(* Logix 5000 project; controller PLC_MCC1300_75F1 vendor 1 type 14 code 166 rev 32.11; software revision 32.04; part 78 of 83 *)
(* tags used below, declared in another part *)
   CM_AreaStackerToLine_JS1_Sync : CM_AreaStackerToLine;
   CM_ConveyorStackerToLine_JS1_Sync : CM_ConveyorStackerToLine;
   M310B : MAC_Conveyor;
   M310B_ALM : MAC_Conveyor_ALM;
   M310B_HMW : MAC_Conveyor_HMW;
   M310Popup : MAC_Popup_ZC[2];
   M311 : MAC_Conveyor;
   M311_ALM : MAC_Conveyor_ALM;
   M311_HMW : MAC_Conveyor_HMW;
   M311A : MAC_Rotator;
   M311A_ALM : MAC_Rotator_ALM;
   M312 : MAC_Conveyor_Single;
   M312_ALM : MAC_Conveyor_ALM;
   M312_HMW : MAC_Conveyor_HMW;
   M350Popup : MAC_Popup_ZC;
   M351 : MAC_Conveyor;
   M351_HMW : MAC_Conveyor_HMW;
   M352 : MAC_Conveyor;
   M352_HMW : MAC_Conveyor_HMW;
   M353 : MAC_Conveyor;
   M353_HMW : MAC_Conveyor_HMW;
   xAlwaysOFF : BOOL;
   xAlwaysON : BOOL;
   Z301 : MAC_Zone_ML;
   Z401 : MAC_Zone;
   Z401_HMR : MAC_Zone_HMR;
   Z401_HMW : MAC_Zone_HMW;
   Z402 : MAC_Zone;
   Z402_ALM : MAC_Zone_ALM;
   Z402_HMR : MAC_Zone_HMR;
   Z402_HMW : MAC_Zone_HMW;
   Z402_INPUT_xMainLineEmergencyON : BOOL;
   Z402_OUTPUT_xMCC_SafetyPanel1 : BOOL;
   Z900 : MAC_Zone;
   Z900_ALM : MAC_Zone_ALM;
   Z900_HMR : MAC_Zone_HMR;
   Z900_HMW : MAC_Zone_HMW;
(* MainProgram, continued *)

   42: [XIC(Z401_HMW.rgxMan.0) OTE(Z401_HMR.rgxMan.0) ,XIC(Z401_HMW.rgxMan.1) OTE(Z401_HMR.rgxMan.1) ];
END_ROUTINE

ROUTINE Z402_Alarm   (* ladder *)
   0: XIC(Z401.tmON_ResetAlarm.DN)FLL(0,Z402_ALM,1);
END_ROUTINE

ROUTINE Z402_Logic   (* ladder *)
   // #####_COSTANTS_#####
   0: NOP();
   // #####_MATCH_#####
   1: NOP();
   // #####_ALARMS_#####
   2: NOP();
   3: XIC(Z402_HMW.xResetErrorRequest)[OTU(Z402_HMW.xResetErrorRequest) ,TOF(Z402.tmON_ResetAlarm,?,?) ];
   4: XIC(Z402.tmON_24Vdc.DN)XIC(Z402.tmON_400Vca.DN)XIC(Z402.tmON_EmergencyOK.DN)OTE(Z402.ST_xEnableControlError);
   5: JSR(Z402_Alarm,0);
   // #####_HMI_LOGICS_#####
   6: NOP();
   // #####_STATUSES_#####
   7: NOP();
   8: [NEQ(Z402_ALM.rgxEmergency[0],0) ,NEQ(Z402_ALM.rgxFault[0],0) ,NEQ(Z402_ALM.rgxWarning[0],0) ,XIC(M310Popup[0].ST_xMachineAlarm) ,XIC(M310Popup[1].ST_xMachineAlarm) ,XIC(M311.ST_xMachineAlarm) ,XIC(M311A.ST_xMachineAlarm) ,XIC(M312.ST_xMachineAlarm) ]OTE(Z402.ST_xZoneError);
   // #####_ZONE MODALITY_#####
   9: NOP();
   // Selector manual mode
   10: XIC(Z402_HMW.xManualModeRequest)OTL(Z402.ST_xSelectionManualMode)OTU(Z402.ST_xSelectionAutomaticMode)OTU(Z402_HMW.xManualModeRequest);
   // Selector automatic mode
   11: XIC(Z402_HMW.xAutomaticModeRequest)OTL(Z402.ST_xSelectionAutomaticMode)OTU(Z402.ST_xSelectionManualMode)OTU(Z402_HMW.xAutomaticModeRequest);
   // Condition Ok for manual mode
   12: [XIC(Z402.ST_xConditionOKStopCycle) ,XIO(Z402.ST_xCycleON) ]OTE(Z402.ST_xConditionOkManualMode);
   // Manual mode accepted
   13: XIC(Z402.ST_xSelectionManualMode)[XIO(Z402.ST_xManualModeAccepted) OTE(Z402.ST_xManualModeRequest) ,[XIC(Z402.ST_xConditionOkManualMode) ,XIC(Z402.ST_xManualModeAccepted) ] OTE(Z402.ST_xManualModeAccepted) ];
   // Auto mode accepted
   14: XIO(Z402.ST_xManualModeAccepted)[XIC(Z402.ST_xSelectionAutomaticMode) ,XIC(Z402.ST_xAutoModeAccepted) ][OTE(Z402.ST_xAutoModeAccepted) ,ONS(Z402.OSR_xAutomaticMode) OTE(Z402.OS_xAutomaticMode) ];
   // Set all manual command for iFix
   15: XIC(Z402.ST_xManualModeAccepted)OTL(M310B_HMW.xEnableDisableManualCommand)OTL(M311_HMW.xEnableDisableManualCommand)OTL(M312_HMW.xEnableDisableManualCommand);
   // Reset all manual command for iFix
   16: XIC(Z402.OS_xAutomaticMode)OTU(M310B_HMW.xEnableDisableManualCommand)OTU(M311_HMW.xEnableDisableManualCommand)OTU(M312_HMW.xEnableDisableManualCommand);
   // #####_LOGICS_#####
   17: NOP();
   18: [XIC(Z402_HMW.xStartCycleRequest) ,XIC(CM_AreaStackerToLine_JS1_Sync.xSB_LineCycle) ]OTE(Z402.OS_xStartCycle);
   19: [XIC(Z402_HMW.xStopCycleRequest) ,XIC(CM_AreaStackerToLine_JS1_Sync.xSB_StopLineCycle) ]OTE(Z402.OS_xStopCycle);
   20: [XIC(Z402.tmON_ForceStop.DN) ONS(Z402.OSR_xForceStopCycle) ,XIC(Z402_HMW.xForceStopCycle) ]OTE(Z402.OS_xForceStopCycle);
   21: XIO(Z402.OS_xForceStopCycle)XIC(Z402.tmON_24Vdc.DN)XIC(Z402.tmON_400Vca.DN)XIC(Z402.tmON_EmergencyOK.DN)OTE(Z402.ST_xConditionOkCycleON);
   22: [XIC(Z402.OS_xStartCycle) ,XIC(Z402.ST_xStartCycleRequest) ]XIC(Z402.ST_xConditionOkCycleON)XIO(Z402.ST_xCycleON)XIO(Z402.OS_xStopCycle)OTE(Z402.ST_xStartCycleRequest);
   23: [XIC(Z402.OS_xStopCycle) ,XIC(Z402.ST_xStopCycleRequest) ]XIC(Z402.ST_xCycleON)XIO(Z402.ST_xStartCycleRequest)OTE(Z402.ST_xStopCycleRequest);
   24: XIC(M310B.ST_xConditionOKStopCycle)XIC(M311.ST_xConditionOKStopCycle)XIC(M311A.ST_xConditionOKStopCycle)XIC(M312.ST_xConditionOKStopCycle)XIC(CM_ConveyorStackerToLine_JS1_Sync.xConditionOkForStopCycle)OTE(Z402.ST_xConditionOKStopCycle);
   25: [XIC(Z402.ST_xStopCycleRequest) XIC(Z402.ST_xConditionOKStopCycle) ,XIC(Z402_HMW.xForceStopCycle) ]OTE(Z402.ST_xStopCycleAccepted);
   // Reimpostare tempo a 15 secondi
   26: [XIC(Z402.ST_xStartCycleRequest) ,XIC(Z402.ST_xCycleON) ]XIC(Z402.ST_xConditionOkCycleON)XIO(Z402.ST_xStopCycleAccepted)XIO(Z402.ST_xManualModeAccepted)[TON(Z402.tmON_Cycle,?,?) ,XIC(Z402.tmON_Cycle.DN) OTE(Z402.ST_xCycleON) ];
   27: XIC(Z402.ST_xCycleON)XIO(Z402.ST_xManualModeRequest)XIO(Z402.ST_xStopCycleRequest)OTE(Z402.ST_xConditionOkPhaseAdvancement);
   28: XIC(Z402.ST_xCycleON)[XIC(M310B.ST_xCleaningAccepted) ,XIO(M310B.ST_xReqCleaning) ][XIC(M311.ST_xCleaningAccepted) ,XIO(M311.ST_xReqCleaning) ][XIC(M312.ST_xCleaningAccepted) ,XIO(M312.ST_xReqCleaning) ]OTE(Z402.ST_xCleaningConditionOK);
   // Speed manager
   29: [MOV(Z402_HMW.dLineSpeed_mm_min,Z402_HMR.dLineSpeed_mm_min) ,LES(Z402_HMR.dLineSpeed_mm_min,35000) MOV(35000,Z402_HMR.dLineSpeed_mm_min) ,GRT(Z402_HMR.dLineSpeed_mm_min,60000) MOV(60000,Z402_HMR.dLineSpeed_mm_min) ];
   // #####_CLEANING_#####
   30: NOP();
   31: XIO(Z402.ST_xCleaningAccepted)XIC(Z402_HMW.xStartCleanZoneRequest)[MOV(Z402_HMW.dCleaningSelection,Z402_HMR.dCleaningSelection) ,OTL(Z402.ST_xReqCleaning) ];
   32: XIC(Z402.ST_xReqCleaning)XIC(Z402.ST_xCleaningConditionOK)[OTL(Z402.ST_xCleaningAccepted) ,OTU(Z402.ST_xReqCleaning) ,OTL(M310B_HMW.xLocalCleaningRequest) ,OTL(M311_HMW.xLocalCleaningRequest) ,OTL(M312_HMW.xLocalCleaningRequest) ];
   33: XIC(Z402_HMW.xStopCleanZoneRequest)[OTU(Z402.ST_xReqCleaning) ,OTU(Z402.ST_xCleaningAccepted) ,MOV(0,Z402_HMW.dCleaningSelection) ,OTU(M310B_HMW.xLocalCleaningRequest) ,OTU(M311_HMW.xLocalCleaningRequest) ,OTU(M311_HMW.xLocalCleaningRequest) ];
   34: XIC(xAlwaysON)[OTU(Z402_HMW.xStartCycleRequest) ,OTU(Z402_HMW.xStopCycleRequest) ,OTU(Z402_HMW.xStartCleanZoneRequest) ,OTU(Z402_HMW.xForceStopCycle) ,OTU(Z402_HMW.xStopCleanZoneRequest) ];
   // #####_HMI_STATUSES_#####
   35: NOP();
   36: XIC(Z402.ST_xZoneError)OTE(Z402_HMR.xZoneAlarm);
   37: [XIC(Z402.ST_xCleaningAccepted) ,XIC(M310B.ST_xCleaningAccepted) XIC(M311.ST_xCleaningAccepted) XIC(M312.ST_xCleaningAccepted) ]OTE(Z402_HMR.xCleaningEnabled);
   38: [MOV(0,Z402_HMR.dCabinetState1) ,[XIC(M310B_ALM.rgxStoppingFault_M[0].1) ,XIC(M311_ALM.rgxStoppingFault_M[0].1) ,XIC(M311A_ALM.rgxStoppingFault_M[0].1) ,XIC(M312_ALM.rgxStoppingFault_M[0].1) ] MOV(2,Z402_HMR.dCabinetState1) ,XIC(Z402_OUTPUT_xMCC_SafetyPanel1) MOV(1,Z402_HMR.dCabinetState1) ];
   39: [XIC(Z402.ST_xManualModeAccepted) MOV(1,Z402_HMR.dZoneMode) ,XIC(Z402.ST_xAutoModeAccepted) MOV(4,Z402_HMR.dZoneMode) ,XIC(Z402.ST_xManualModeRequest) MOV(8,Z402_HMR.dZoneMode) ];
   40: [MOV(2,Z402_HMR.dZoneState) ,XIC(Z402.ST_xStartCycleRequest) XIO(Z402.ST_xCycleON) MOV(4,Z402_HMR.dZoneState) ,XIC(Z402.ST_xCycleON) MOV(1,Z402_HMR.dZoneState) ,XIC(Z402.ST_xStopCycleRequest) MOV(8,Z402_HMR.dZoneState) ,XIO(Z402_INPUT_xMainLineEmergencyON) MOV(1024,Z402_HMR.dZoneState) ];
   41: [[XIC(Z402.ST_xCleaningAccepted) ,XIC(M310B.ST_xCleaningAccepted) XIC(M311.ST_xCleaningAccepted) XIC(M312.ST_xCleaningAccepted) ] MOV(1,Z402_HMR.dCleaningState) ,XIO(Z402.ST_xCleaningAccepted) MOV(2,Z402_HMR.dCleaningState) ,XIC(Z402.ST_xReqCleaning) XIO(Z402.ST_xCleaningAccepted) MOV(4,Z402_HMR.dCleaningState) ];
   42: [XIC(Z402_HMW.rgxMan.0) OTE(Z402_HMR.rgxMan.0) ,XIC(Z402_HMW.rgxMan.1) OTE(Z402_HMR.rgxMan.1) ];
END_ROUTINE

ROUTINE Z900_Alarm   (* ladder *)
   0: XIC(Z900.tmON_ResetAlarm.DN)FLL(0,Z900_ALM,1);
END_ROUTINE

ROUTINE Z900_Logic   (* ladder *)
   // #####_COSTANTS_#####
   0: NOP();
   // #####_MATCH_#####
   1: NOP();
   2: XIC(Z301.INPUT_x24VdcVoltageON)XIC(Z301.INPUT_xPowerSupply24VLogic1)XIC(Z301.INPUT_xPowerSupply24VLogic2)XIC(Z301.INPUT_xPowerSupply24VLogic3)XIC(Z301.INPUT_xEthernetSwitch24VON)XIC(Z301.INPUT_xPowerSupply24VDrive1)XIC(Z301.INPUT_xPowerSupply24VDrive2)TON(Z900.tmON_24Vdc,?,?);
   3: XIC(Z301.INPUT_xPowerSupply400VDrive1)XIC(Z301.INPUT_xPowerSupply400VDrive2)TON(Z900.tmON_400Vca,?,?);
   4: XIC(Z301.INPUT_xMainEmergencyON)TON(Z900.tmON_EmergencyOK,?,?);
   // #####_ALARMS_#####
   5: NOP();
   6: XIC(Z900_HMW.xResetErrorRequest)[OTU(Z900_HMW.xResetErrorRequest) ,TOF(Z900.tmON_ResetAlarm,?,?) ];
   7: XIC(Z900.tmON_24Vdc.DN)XIC(Z900.tmON_400Vca.DN)XIC(Z900.tmON_EmergencyOK.DN)OTE(Z900.ST_xEnableControlError);
   8: JSR(Z900_Alarm,0);
   // #####_HMI_LOGICS_#####
   9: NOP();
   // #####_STATUSES_#####
   10: NOP();
   11: [NEQ(Z900_ALM.rgxEmergency[0],0) ,NEQ(Z900_ALM.rgxFault[0],0) ,NEQ(Z900_ALM.rgxWarning[0],0) ,XIC(M351.ST_xMachineAlarm) ,XIC(M352.ST_xMachineAlarm) ,XIC(M353.ST_xMachineAlarm) ]OTE(Z900.ST_xZoneError);
   // #####_ZONE MODALITY_#####
   12: NOP();
   // Selector manual mode
   13: XIC(Z900_HMW.xManualModeRequest)OTL(Z900.ST_xSelectionManualMode)OTU(Z900.ST_xSelectionAutomaticMode)OTU(Z900_HMW.xManualModeRequest);
   // Selector automatic mode
   14: XIC(Z900_HMW.xAutomaticModeRequest)OTL(Z900.ST_xSelectionAutomaticMode)OTU(Z900.ST_xSelectionManualMode)OTU(Z900_HMW.xAutomaticModeRequest);
   // Condition Ok for manual mode
   15: [XIC(Z900.ST_xConditionOKStopCycle) ,XIO(Z900.ST_xCycleON) ]OTE(Z900.ST_xConditionOkManualMode);
   // Manual mode accepted
   16: XIC(Z900.ST_xSelectionManualMode)[XIO(Z900.ST_xManualModeAccepted) OTE(Z900.ST_xManualModeRequest) ,[XIC(Z900.ST_xConditionOkManualMode) ,XIC(Z900.ST_xManualModeAccepted) ] OTE(Z900.ST_xManualModeAccepted) ];
   // Auto mode accepted
   17: XIO(Z900.ST_xManualModeAccepted)[XIC(Z900.ST_xSelectionAutomaticMode) ,XIC(Z900.ST_xAutoModeAccepted) ][OTE(Z900.ST_xAutoModeAccepted) ,ONS(Z900.OSR_xAutomaticMode) OTE(Z900.OS_xAutomaticMode) ];
   // Set all manual command for iFix
   18: XIC(Z900.ST_xManualModeAccepted)OTL(M351_HMW.xEnableDisableManualCommand)OTL(M352_HMW.xEnableDisableManualCommand)OTL(M353_HMW.xEnableDisableManualCommand);
   // Reset all manual command for iFix
   19: XIC(Z900.OS_xAutomaticMode)OTU(M351_HMW.xEnableDisableManualCommand)OTU(M352_HMW.xEnableDisableManualCommand)OTU(M353_HMW.xEnableDisableManualCommand);
   20: XIO(M350Popup.INPUT_xPopupHigh)OTU(M351_HMW.xEnableDisableManualCommand);
   // #####_LOGICS_#####
   21: NOP();
   22: XIC(Z900_HMW.xStartCycleRequest)OTE(Z900.OS_xStartCycle);
   23: XIC(Z900_HMW.xStopCycleRequest)OTE(Z900.OS_xStopCycle);
   24: XIC(xAlwaysOFF)TON(Z900.tmON_ForceStop,?,?);
   25: [XIC(Z900.tmON_ForceStop.DN) ONS(Z900.OSR_xForceStopCycle) ,XIC(Z900_HMW.xForceStopCycle) ]OTE(Z900.OS_xForceStopCycle);
   26: XIO(Z900.OS_xForceStopCycle)XIC(Z900.tmON_24Vdc.DN)XIC(Z900.tmON_400Vca.DN)XIC(Z900.tmON_EmergencyOK.DN)XIO(Z900.ST_xManualModeAccepted)OTE(Z900.ST_xConditionOkCycleON);
   27: [XIC(Z900.OS_xStartCycle) ,XIC(Z900.ST_xStartCycleRequest) ]XIC(Z900.ST_xConditionOkCycleON)[XIO(Z900.ST_xCycleON) ,XIC(Z900.ST_xStopCycleRequest) ]XIO(Z900.OS_xStopCycle)OTE(Z900.ST_xStartCycleRequest);
   28: [XIC(Z900.OS_xStopCycle) ,XIC(Z900.ST_xStopCycleRequest) ]XIC(Z900.ST_xCycleON)XIO(Z900.ST_xStartCycleRequest)OTE(Z900.ST_xStopCycleRequest);
   29: XIC(M351.ST_xConditionOKStopCycle)XIC(M352.ST_xConditionOKStopCycle)XIC(M353.ST_xConditionOKStopCycle)OTE(Z900.ST_xConditionOKStopCycle);
   30: [XIC(Z900.ST_xStopCycleRequest) XIC(Z900.ST_xConditionOKStopCycle) ,XIC(Z900_HMW.xForceStopCycle) ]OTE(Z900.ST_xStopCycleAccepted);
   // Rimettere il timer a 15s
   31: [XIC(Z900.ST_xStartCycleRequest) ,XIC(Z900.ST_xCycleON) ]XIC(Z900.ST_xConditionOkCycleON)XIO(Z900.ST_xStopCycleAccepted)[TON(Z900.tmON_Cycle,?,?) ,XIC(Z900.tmON_Cycle.DN) OTE(Z900.ST_xCycleON) ];
   32: XIC(Z900.ST_xCycleON)XIO(Z900.ST_xManualModeRequest)XIO(Z900.ST_xStopCycleRequest)OTE(Z900.ST_xConditionOkPhaseAdvancement);
   // Speed manager
   33: [MOV(Z900_HMW.dLineSpeed_mm_min,Z900_HMR.dLineSpeed_mm_min) ,LES(Z900_HMR.dLineSpeed_mm_min,35000) MOV(35000,Z900_HMR.dLineSpeed_mm_min) ,GRT(Z900_HMR.dLineSpeed_mm_min,90000) MOV(90000,Z900_HMR.dLineSpeed_mm_min) ];
   34: XIC(Z900.ST_xCycleON)[XIC(M351.ST_xCleaningAccepted) ,GRT(Z900_HMW.dCleaningSelection,3510) ][XIC(M352.ST_xCleaningAccepted) ,GRT(Z900_HMW.dCleaningSelection,3520) ][XIC(M353.ST_xCleaningAccepted) ,GRT(Z900_HMW.dCleaningSelection,3530) ]OTE(Z900.ST_xCleaningConditionOK);
   // #####_CREANING_#####
   35: NOP();
   36: XIO(Z900.ST_xCleaningAccepted)XIC(Z900_HMW.xStartCleanZoneRequest)[MOV(Z900_HMW.dCleaningSelection,Z900_HMR.dCleaningSelection) ,OTL(Z900.ST_xReqCleaning) ];
   37: XIC(Z900.ST_xReqCleaning)XIC(Z900.ST_xCleaningConditionOK)[OTL(Z900.ST_xCleaningAccepted) ,OTU(Z900.ST_xReqCleaning) ];
   38: XIC(Z900_HMW.xStopCleanZoneRequest)[OTU(Z900.ST_xReqCleaning) ,OTU(Z900.ST_xCleaningAccepted) ,MOV(0,Z900_HMW.dCleaningSelection) ,OTU(M351_HMW.xLocalCleaningRequest) ,OTU(M352_HMW.xLocalCleaningRequest) ,OTU(M352_HMW.xLocalCleaningRequest) ];
   39: XIC(xAlwaysON)[OTU(Z900_HMW.xStartCycleRequest) ,OTU(Z900_HMW.xStopCycleRequest) ,OTU(Z900_HMW.xStartCleanZoneRequest) ,OTU(Z900_HMW.xForceStopCycle) ,OTU(Z900_HMW.xStopCleanZoneRequest) ];
